// TIA Portal project "S7_1516_LECTOR620_DI" (V15)

(* hardware
DEVICE "S71500/ET200MP station_1"  S7-1500 station
   slot 0: "Rail_0"  Rack  6ES7 590-1***0-0AA0
   slot 0: "PM 190W 120/230VAC"  PM 190W 120/230VAC  6EP1333-4BA00
   slot 1: "PLC_1"  CPU 1516-3 PN/DP  6ES7 516-3AN00-0AB0  V1.8
      slot 3: "CPU display_1"  6ES7591-1BA00-0AA0
   slot 2: "DI 32x24VDC HF_1"  DI 32x24VDC HF  6ES7 521-1BL00-0AB0  V2.1
   slot 3: "DQ 32x24VDC/0.5A ST_1"  DQ 32x24VDC/0.5A ST  6ES7 522-1BL00-0AB0  V2.0
   slot 4: "AI 8xU/I/RTD/TC ST_1"  AI 8xU/I/RTD/TC ST  6ES7 531-7KF00-0AB0  V2.0
   slot 5: "AQ 4xU/I ST_1"  AQ 4xU/I ST  6ES7 532-5HD00-0AB0  V2.0
DEVICE "HMI_1"  TP700 Comfort
   slot 0: "HMI_1"  TP700 Comfort  6AV2 124-0GC01-0AX0  15.0.0.0
   slot 1: "HMI_RT_1"  TP700 Comfort  6AV2 124-0GC01-0AX0  15.0.0.0
   slot 5: "HMI_1.IE_CP_1"  PROFINET Interface  15.0.0.0
      slot 1: "PROFINET Interface_1"  PROFINET Interface
         slot 1: "Port_1"  Port
         slot 2: "Port_2"  Port
   slot 7: "HMI_1.MPI/DP_CP_1"  MPI/DP Interface  15.0.0.0
DEVICE "GSD device_2"  GSD.Device.PN
   slot 0: "Rack"  Rack  V1.0
   slot 0: "LECTOR62x"  LECTOR62x  HandShake (HS)  V1.1.0
      slot 0: "LECTOR62x  HandShake (HS)"  LECTOR62x  HandShake (HS)
      slot 1: "Interface"  Interface
         slot 1: "Port 1"  Port 1
   slot 1: "Ctrl Bits in_1"  Ctrl Bits in
      slot 0: "Ctrl Bits in"  Ctrl Bits in
   slot 2: "Ctrl Bits out_1"  Ctrl Bits out
      slot 0: "Ctrl Bits out"  Ctrl Bits out
   slot 3: " 32 Byte Input (HS)_1"   32 Byte Input (HS)
      slot 0: " 32 Byte Input (HS)"   32 Byte Input (HS)
   slot 4: " 32 Byte Output (HS)_1"   32 Byte Output (HS)
      slot 0: " 32 Byte Output (HS)"   32 Byte Output (HS)
DEVICE "PC-System_1"  SIMATIC PC station
   slot 0: "SIMATIC PC station"  Rail  SIMATIC PC-Station  V1.0
      slot 125: "Stationmanager"  Station_Manager  V6.0.4
   slot 1: "IE general_1"  IE General  IE_CP  V8.2.0
   slot 3: "HMI_RT_2"  WinCC RT Advanced  6AV2 104-0xxxx-xxxx  15.0.0.0
      slot 33792: "Host interface"  Host interface
*)

// ===== PLC "PLC_1"  CPU 1516-3 PN/DP =====

VAR_GLOBAL   // PLC tag table "Default tag table"
   "AD_CH0" AT %IW4 : Int;
   "Sensor1" AT %I0.0 : Bool;
   "Tag_5" AT %IW58 : Int;
   "Tag_6" AT %IW12 : Int;
   "DA_CH0" AT %QW4 : Int;
   "SICK_IN_1" AT %Q0.0 : Bool;
   "Tag_3" AT %Q0.1 : Bool;
   "Tag_4" AT %QW1 : Int;
   "Tag_7" AT %Q0.2 : Bool;
   "Tag_8" AT %Q1.1 : Bool;
   "Tag_9" AT %Q1.2 : Bool;
   "Clock_Byte" AT %MB0 : Byte;
   "Clock_10Hz" AT %M0.0 : Bool;
   "Clock_5Hz" AT %M0.1 : Bool;
   "Clock_2.5Hz" AT %M0.2 : Bool;
   "Clock_2Hz" AT %M0.3 : Bool;
   "Clock_1.25Hz" AT %M0.4 : Bool;
   "Clock_1Hz" AT %M0.5 : Bool;
   "Clock_0.625Hz" AT %M0.6 : Bool;
   "Clock_0.5Hz" AT %M0.7 : Bool;
   "SignalUlaz" AT %M1.0 : Bool;
   "SICK_OUT_1" AT %I0.1 : Bool;
   "SICK_OUT_1_MEM" AT %M10.0 : Bool;
   "Tag_1" AT %M100.0 : Bool;
   "Tag_2" AT %M100.1 : Bool;
   "Tag_10" AT %M100.2 : Bool;
   "Tag_11" AT %M100.3 : Bool;
   "Tag_12" AT %MW101 : Word;
   "Request" AT %M100.4 : Bool;
   "No_of_counts_in" AT %IB57 : Byte;
   "No_of_counts_out" AT %QB49 : Byte;
   "SICK_OUT_1_old" AT %M2.0 : Bool;
   "Code_byte_1" AT %IB62 : Byte;
   "Tag_13" AT %MW3 : Int;
   "MOVE_ERROR" AT %MW4 : Int;
   "Tag_14" AT %IB56 : Byte;
   "Code_byte_2" AT %IB63 : Char;
   "Code_byte_3" AT %IB64 : Char;
   "Code_byte_4" AT %IB65 : Char;
   "Code_byte_5" AT %IB66 : Char;
   "Code_byte_6" AT %IB67 : Char;
   "Code_byte_7" AT %IB68 : Char;
   "Code_byte_8" AT %IB69 : Char;
   "Code_byte_9" AT %IB70 : Char;
   "Code_byte_10" AT %IB71 : Char;
   "Code_byte_11" AT %IB72 : Char;
   "Code_byte_12" AT %IB73 : Char;
   "Code_byte_13" AT %IB74 : Char;
   "ADDA_ENABLE" AT %I0.2 : Bool;
   "DA_CH2" AT %QW8 : Int;
   "AD_CH2" AT %IW8 : Int;
   "AD_CH1" AT %IW6 : Int;
   "AD_CH3" AT %IW10 : Int;
   "DA_CH1" AT %QW6 : Int;
   "DA_CH3" AT %QW10 : Int;
   "iCounter_Tag_kopija" AT %QW12 : Int;
   "PrebranaKoda" AT %QW14 : WChar;
   "Tag_15" AT %I0.3 : Bool;
   "Tag_16" AT %Q0.3 : Bool;
   "Tag_17" AT %Q2.0 : Bool;
   "Tag_18" AT %Q2.1 : Bool;
   "Tag_19" AT %Q2.2 : Bool;
END_VAR

// folder: SICK AG

TYPE "ST_SICK_Lector_CLV6xx"
TITLE = SICK Lector/CLV6xx data type
VERSION : 0.1
// This data type includes arguments and results using by the SICK_Lector_CLV6xx_PNDP function block.
   STRUCT
      Matchcode : Struct   // ==Matchcode==
         sName : String[10];   // Matchcode number (Match[1..9]) (Input)
         nCodeType : Char;   // Code type see device documentation. (Example: 'd'= EAN-Code; 's'=QR-Code; '*'= Don't care) (Input)
         iMinMaxLength : USInt;   // Sets the min and may length. 0= Don't care (Input)
         sContent : String[75];   // Matchcode content
      END_STRUCT;
      FreeCommand : Struct   // ==Free Command==
         sCommand : String[100];   // Command (SICK CoLa-A protocol without [STX]/[ETX] framing) (In)
         sResult : String[100];   // Result (SICK CoLa-A protocol) (Out)
      END_STRUCT;
      ReadingResult : Struct   // ==Reading Result==
         iCounter : USInt;   // This counter is incremented if a new reading result has arrived (In)
         iLength : Int;   // Byte length of the reading result (Out)
         arrResult : Array[1..200] of Byte;   // Reading result data defined in the SOPAS output format (Out)
      END_STRUCT;
   END_STRUCT;
END_TYPE

// folder: (top level)

DATA_BLOCK "Data_block_1"   // DB1
{ S7_Optimized_Access := 'FALSE' }
VERSION : 0.1
   VAR
      Error_Detektovan : Bool;   // 1 ce je prislo do napake
      Error_Koda : DWord;   // ID koda napake
      startFound : Bool;   // za Move_Code funkcijo
      endFound : Bool;   // za Move_Code funkcijo
      Sensor_ok_blink : Byte;
      No_of_counts : LInt;
      DA0 : Real;
      AD0 : Real;
      DA2 : Real;
      AD2 : Real;
      Static_1 : Array[0..5] of Int;
      TestBitStefanRequest : Bool;
      ShranjenaPrebranaKoda_Cas : Date_And_Time := DT#2021-05-14-08:00:42.263;
      ShranjenaPrebranaKoda : String;
      Operand1 : Bool;
      DatumInCas : Struct
         Datum : Bool;
         Ura : Bool;
      END_STRUCT;
      AD3 : Real;
      Prebrana_Koda_FLAG : Bool;
      Counter_1_Reset : Bool;
      Operand2 : Bool;
   END_VAR
BEGIN
END_DATA_BLOCK

DATA_BLOCK "IDB_Lector6xx"   // DB2
{ S7_Optimized_Access := 'TRUE' }
AUTHOR : SICKAG
FAMILY : Ident
VERSION : 1.2
// stored: InstanceOfName SICK_Lector_CLV6xx_PNDP
"SICK_Lector_CLV6xx_PNDP"
BEGIN
END_DATA_BLOCK

DATA_BLOCK "DB_Example"   // DB3
{ S7_Optimized_Access := 'TRUE' }
VERSION : 0.1
   VAR
      stEdge : Struct   // Edge detection flags
         xEdgeTrigger : Bool;
         xEdgeMatchcode : Bool;
         xEdgeDone : Bool;
         xEdgeError : Bool;
         xEdgeTriggerMem : Bool;
         xEdgeDoneMem : Bool;
         xEdgeErrorMem : Bool;
         xEdgeMatchcodeMem : Bool;
      END_STRUCT;
      xTrigger : Bool;   // Start read tag command
      xMatchcode : Bool;
      xTriggerDone : Bool;   // Read tag done
      xMatchcodeDone : Bool;
      sReadingResult : String[200];   // Read content
      stLector : "ST_SICK_Lector_CLV6xx";   // RFU data
      arrReadingResult : Array[0..199] of Byte;   // Read content backup
   END_VAR
BEGIN
END_DATA_BLOCK

DATA_BLOCK "SICK_Lector_CLV6xx_PNDP_DB"   // DB4
{ S7_Optimized_Access := 'TRUE' }
AUTHOR : SICKAG
FAMILY : Ident
VERSION : 1.2
// stored: InstanceOfName SICK_Lector_CLV6xx_PNDP
"SICK_Lector_CLV6xx_PNDP"
BEGIN
END_DATA_BLOCK

DATA_BLOCK "Block_1_DB"   // DB5
{ S7_Optimized_Access := 'TRUE' }
AUTHOR : Stefan_Milivojcev
VERSION : 0.1
// stored: InstanceOfName Block_1
"Block_1"
BEGIN
END_DATA_BLOCK

// folder: System blocks/Program resources

DATA_BLOCK "IEC_Counter_0_DB"   // DB6
{ S7_Optimized_Access := 'TRUE' }
AUTHOR : SIMATIC
FAMILY : IEC
NAME : LCNTR
VERSION : 1.2
// stored: InstanceOfName IEC_LCOUNTER
"IEC_LCOUNTER"
BEGIN
END_DATA_BLOCK

// folder: (top level)

FUNCTION_BLOCK "Block_1"   // FB1, SCL
TITLE = Shranjevanje_Branja
{ S7_Optimized_Access := 'TRUE' }
AUTHOR : Stefan_Milivojcev
VERSION : 0.1
   VAR_INPUT
      RESULT_ARRAY_SIZE : Int;   // Velikost najvecjega moznega rezultata branja
      Date_Time_Temp : Date_And_Time;
   END_VAR
   VAR_OUTPUT
      startFound : Bool;
      endFound : Bool;
      PrebranaKoda_Cas : Date_And_Time;
      PrebranaKoda : String;
   END_VAR
   VAR_TEMP
      i : Int;
   END_VAR
BEGIN
   //Stefan Milivojčev
   //stefan.milivojcev@gmail.com
   //
   //Prepoznava START in STOP bita


   #startFound := FALSE;
   #endFound := FALSE;
   #i := 0;
   #PrebranaKoda := '';



   IF ("DB_Example".stLector.ReadingResult.arrResult[1] = 16#02) THEN
       // Statement section IF
       #startFound := 1;
   END_IF;

   IF (#startFound = 1) THEN //ce smo najdli zacetek kode iscemo konec

       FOR #i := 1 TO #RESULT_ARRAY_SIZE DO
           // Statement section FOR

           IF ("DB_Example".stLector.ReadingResult.arrResult[#i] = 16#03) THEN
               // Statement section IF
               #endFound := TRUE;

           ELSE

               #PrebranaKoda[#i - 1] := "DB_Example".stLector.ReadingResult.arrResult[#i];

           END_IF;



       END_FOR;

       #PrebranaKoda_Cas := #Date_Time_Temp;


   END_IF;




   "Data_block_1".No_of_counts := "DB_Example".stLector.ReadingResult.iCounter;
END_FUNCTION_BLOCK

ORGANIZATION_BLOCK "Main"   // OB1, LAD, ProgramCycle
TITLE = "Main Program Sweep (Cycle)"
{ S7_Optimized_Access := 'TRUE' }
VERSION : 0.1
   VAR_INPUT
      Initial_Call : Bool;   // Initial call of this OB
      Remanence : Bool;   // =True, if remanent data are available
   END_VAR
   VAR_TEMP
      Temp_3 : Real;
      Temp_2 : LInt;
      Temp_Cas_Branja : Date_And_Time;
      Temp3 : Date;
      Temp4 : DInt;
      temp6 : Bool;
      Temp5 : UInt;
   END_VAR
   VAR_TEMP   // added for the SCL form of the ladder/FBD networks
      _w1 : Bool;
      _w2 : Bool;
   END_VAR
BEGIN

REGION Network 1: Request za branje
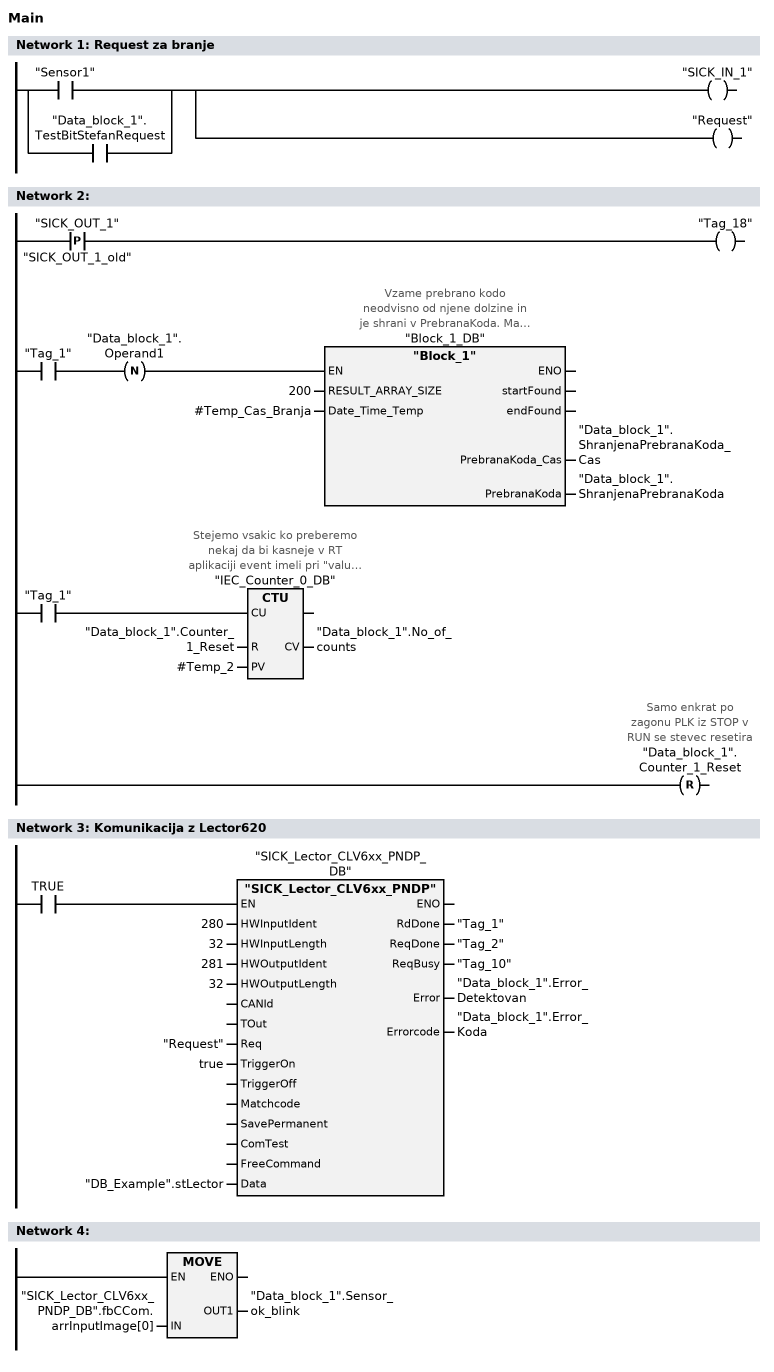
   RUNG wire#powerrail
      Contact( "Sensor1" )
      wire#w1
      Coil( "SICK_IN_1" )
   END_RUNG
   RUNG wire#powerrail
      Contact( "Data_block_1".TestBitStefanRequest )
   END_RUNG wire#w1
   RUNG wire#w1
      Coil( "Request" )
   END_RUNG
   // the same network as SCL:
   "SICK_IN_1" := "Sensor1" OR "Data_block_1".TestBitStefanRequest;
   "Request" := "SICK_IN_1";
END_REGION

REGION Network 2
   #_w1 := "SICK_OUT_1" AND NOT "SICK_OUT_1_old";   // rising edge of "SICK_OUT_1"
   "SICK_OUT_1_old" := "SICK_OUT_1";
   "Tag_18" := #_w1;
   #_w2 := NOT "Tag_1" AND "Data_block_1".Operand1;   // falling edge
   "Data_block_1".Operand1 := "Tag_1";
   IF #_w2 THEN
       "Block_1_DB"(RESULT_ARRAY_SIZE := 200,   // "Block_1": Vzame prebrano kodo neodvisno od njene dolzine in je shrani v PrebranaKoda. Max dolzina je trenutno 200
                    Date_Time_Temp := #Temp_Cas_Branja,
                    PrebranaKoda_Cas => "Data_block_1".ShranjenaPrebranaKoda_Cas,
                    PrebranaKoda => "Data_block_1".ShranjenaPrebranaKoda);
   END_IF;
   "IEC_Counter_0_DB".CTU(CU := "Tag_1",   // Stejemo vsakic ko preberemo nekaj da bi kasneje v RT aplikaciji event imeli pri "value change"
                          R := "Data_block_1".Counter_1_Reset,
                          PV := #Temp_2,
                          CV => "Data_block_1".No_of_counts);
   "Data_block_1".Counter_1_Reset := FALSE;   // Samo enkrat po zagonu PLK iz STOP v RUN se stevec resetira
END_REGION

REGION Network 3: Komunikacija z Lector620
   RUNG wire#powerrail
      Contact( TRUE )
      "SICK_Lector_CLV6xx_PNDP_DB"(HWInputIdent := 280, HWInputLength := 32, HWOutputIdent := 281, HWOutputLength := 32, CANId :=, TOut :=, Req := "Request", TriggerOn := true, TriggerOff :=, Matchcode :=, SavePermanent :=, ComTest :=, FreeCommand :=, Data := "DB_Example".stLector, RdDone => "Tag_1", ReqDone => "Tag_2", ReqBusy => "Tag_10", Error => "Data_block_1".Error_Detektovan, Errorcode => "Data_block_1".Error_Koda)
   END_RUNG
   // the same network as SCL:
   IF TRUE THEN
       "SICK_Lector_CLV6xx_PNDP_DB"(HWInputIdent := 280,   // "SICK_Lector_CLV6xx_PNDP"
                               HWInputLength := 32,
                               HWOutputIdent := 281,
                               HWOutputLength := 32,
                               Req := "Request",
                               TriggerOn := true,
                               Data := "DB_Example".stLector,
                               RdDone => "Tag_1",
                               ReqDone => "Tag_2",
                               ReqBusy => "Tag_10",
                               Error => "Data_block_1".Error_Detektovan,
                               Errorcode => "Data_block_1".Error_Koda);
   END_IF;
END_REGION

REGION Network 4
   RUNG wire#powerrail
      Move(in := "SICK_Lector_CLV6xx_PNDP_DB".fbCCom.arrInputImage[0], out1 => "Data_block_1".Sensor_ok_blink)
   END_RUNG
   // the same network as SCL:
   "Data_block_1".Sensor_ok_blink := "SICK_Lector_CLV6xx_PNDP_DB".fbCCom.arrInputImage[0];
END_REGION
END_ORGANIZATION_BLOCK

ORGANIZATION_BLOCK "Cyclic interrupt"   // OB30, LAD, CyclicInterrupt
{ S7_Optimized_Access := 'TRUE' }
VERSION : 0.1
   VAR_INPUT
      Initial_Call : Bool;   // Initial call of this OB
      Event_Count : Int;   // Events discarded
   END_VAR
BEGIN

REGION Network 1
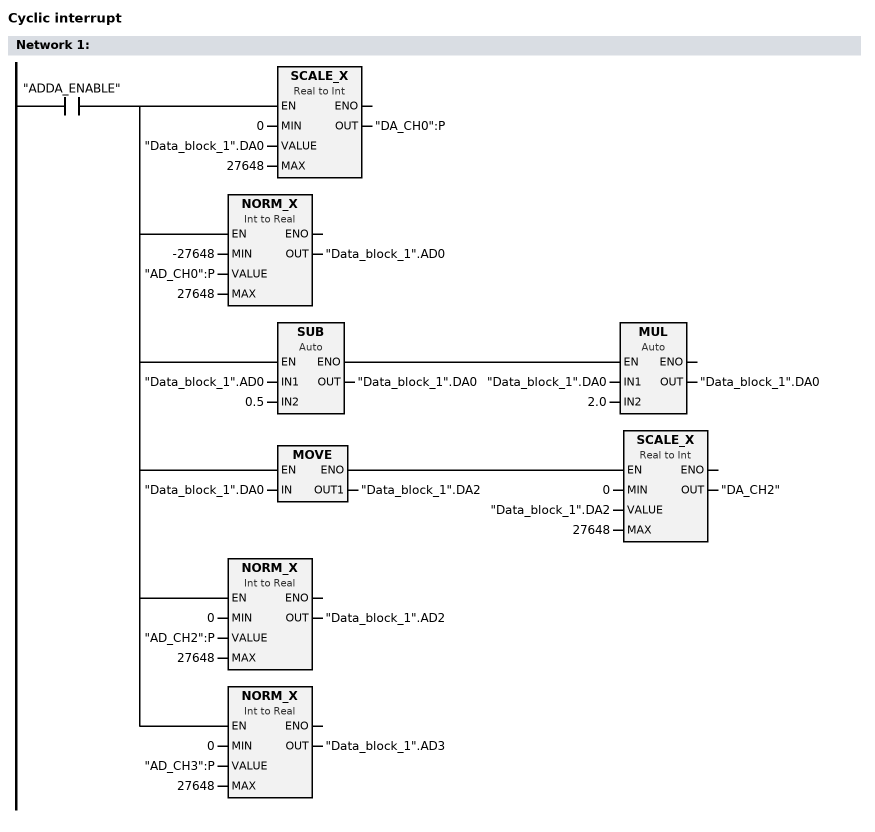
   RUNG wire#powerrail
      Contact( "ADDA_ENABLE" )
      wire#w1
      { S7_Templates := "[SrcType := Real, DestType := Int]" } Scale(min := 0, value := "Data_block_1".DA0, max := 27648, out => "DA_CH0":P)
   END_RUNG
   RUNG wire#w1
      { S7_Templates := "[SrcType := Int, DestType := Real]" } Normalize(min := -27648, value := "AD_CH0":P, max := 27648, out => "Data_block_1".AD0)
   END_RUNG
   RUNG wire#w1
      Sub(in1 := "Data_block_1".AD0, in2 := 0.5, out => "Data_block_1".DA0)
      Mul(in1 := "Data_block_1".DA0, in2 := 2.0, out => "Data_block_1".DA0)
   END_RUNG
   RUNG wire#w1
      Move(in := "Data_block_1".DA0, out1 => "Data_block_1".DA2)
      { S7_Templates := "[SrcType := Real, DestType := Int]" } Scale(min := 0, value := "Data_block_1".DA2, max := 27648, out => "DA_CH2")
   END_RUNG
   RUNG wire#w1
      { S7_Templates := "[SrcType := Int, DestType := Real]" } Normalize(min := 0, value := "AD_CH2":P, max := 27648, out => "Data_block_1".AD2)
   END_RUNG
   RUNG wire#w1
      { S7_Templates := "[SrcType := Int, DestType := Real]" } Normalize(min := 0, value := "AD_CH3":P, max := 27648, out => "Data_block_1".AD3)
   END_RUNG
   // the same network as SCL:
   IF "ADDA_ENABLE" THEN
       "DA_CH0":P := SCALE_X(MIN := 0, VALUE := "Data_block_1".DA0, MAX := 27648);
       "Data_block_1".AD0 := NORM_X(MIN := -27648, VALUE := "AD_CH0":P, MAX := 27648);
       "Data_block_1".DA0 := "Data_block_1".AD0 - 0.5;
       "Data_block_1".DA0 := "Data_block_1".DA0 * 2.0;
       "Data_block_1".DA2 := "Data_block_1".DA0;
       "DA_CH2" := SCALE_X(MIN := 0, VALUE := "Data_block_1".DA2, MAX := 27648);
       "Data_block_1".AD2 := NORM_X(MIN := 0, VALUE := "AD_CH2":P, MAX := 27648);
       "Data_block_1".AD3 := NORM_X(MIN := 0, VALUE := "AD_CH3":P, MAX := 27648);
   END_IF;
END_REGION
END_ORGANIZATION_BLOCK

ORGANIZATION_BLOCK "Startup"   // OB100, LAD, Startup
TITLE = "Complete Restart"
{ S7_Optimized_Access := 'TRUE' }
VERSION : 0.1
   VAR_INPUT
      LostRetentive : Bool;   // True if retentive data are lost
      LostRTC : Bool;   // True if date and time are lost
   END_VAR
   VAR_TEMP
      operand1 : Bool;
   END_VAR
BEGIN

REGION Network 1
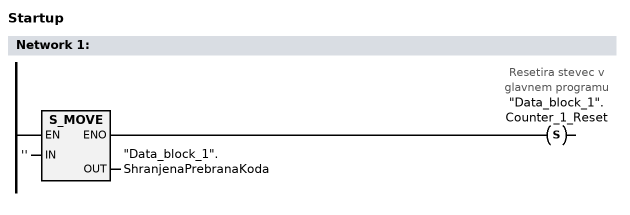
   RUNG wire#powerrail
      S_Move(in := '', out => "Data_block_1".ShranjenaPrebranaKoda)
      S_Coil( "Data_block_1".Counter_1_Reset )   // Resetira stevec v glavnem programu
   END_RUNG
   // the same network as SCL:
   "Data_block_1".ShranjenaPrebranaKoda := '';
   "Data_block_1".Counter_1_Reset := TRUE;   // Resetira stevec v glavnem programu
END_REGION
END_ORGANIZATION_BLOCK

// folder: SICK AG

FUNCTION_BLOCK "SICK_Lector_CLV6xx_PNDP"   // FB72, SCL
TITLE = SICK Lector6xx / CLV6xx function block
{ S7_Optimized_Access := 'TRUE' }
AUTHOR : SICKAG
FAMILY : Ident
VERSION : 1.2
// This function block is used for a communication between a SICK Lector6xx / SICK CLV6xx code reader and a Siemens S7-1200/S7-1500 PLC via  PROFINET/PROFIBUS
   VAR_INPUT
      HWInputIdent : Hw_Io;   // Hardware identification number of the input module
      HWInputLength : USInt;   // Size of the input module
      HWOutputIdent : Hw_Io;   // Hardware identification number of the output module
      HWOutputLength : USInt;   // Size of the output module
      CANId : USInt;   // CAN ID (0= Master / No CAN network)
      TOut : Time := T#10s;   // Time out
      Req : Bool;   // A positive edge starts the request
      TriggerOn : Bool;   // Select: Trigger On to open the reading gate via a SW-Trigger command
      TriggerOff : Bool;   // Select: Trigger Off to close the reading gate via a SW-Trigger command
      Matchcode : Bool;   // Select: Matchcode (details at #Data)
      SavePermanent : Bool;   // Select: Save permanent
      ComTest : Bool;   // Select: Communication test
      FreeCommand : Bool;   // Select: Free command (details at #Data)
   END_VAR
   VAR_OUTPUT
      RdDone : Bool;   // Positive edge: A reading result sent by the device was received
      ReqDone : Bool;   // Request done / Indicates whether a CoLa command was sent and an answer was received
      ReqBusy : Bool;   // Request in process / Request processing
      Error : Bool;   // Error detected
      Errorcode : DWord;   // Error code (see documentation)
   END_VAR
   VAR_IN_OUT
      Data : "ST_SICK_Lector_CLV6xx";   // Command arguments and result outputs of the FB actions
   END_VAR
   VAR
      bTriggerReq : Bool;   // Rising edge detection
      bTriggerReqMem : Bool;   // Rising edge detection
      bTriggerDone : Bool;   // Rising edge detection
      bTriggerDoneMem : Bool;   // Rising edge detection
      bTriggerError : Bool;   // Rising edge detection
      bTriggerErrorMem : Bool;   // Rising edge detection
      bCanActive : Bool;   // CAN-Bus active flag
      bDeviceState : Bool;   // Current device state (True= Edit-Mode | False= Run-Mode)
      bEnforceLogout : Bool;   // Logout enforced
      bReqBusyMem : Bool;   // Backup variable
      iStep : USInt;   // Currrent FB step
      iCommandIndex : Int;   // Command index
      iCommandLength : UInt;   // Length of the command that should be send
      iRecordSize : UInt;   // Length of the record array
      iCommandSize : UInt;   // Length of the command array
      iReadingResultSize : UInt;   // Length of the reading result array
      iIndex : UInt;   // Index variable
      nTempErrorCode : DWord;   // Temporarily error code
      nLogoutErrorCode : DWord;   // Temporarily error code
      arrSelection : Array[0..5] of Bool;   // input bit selection
      arrCommand : Array[0..499] of Byte;   // Contains the transmitted CoLa command
      arrRecord : Array[0..499] of Byte;   // Contains the received telegram
      fbTimeout : TON_TIME;   // Instance: Timer on delay (Time out)
      fbCCom : "SICK_CCOMM_PNDP";   // Instance: CoLa communication block
   END_VAR
   VAR_TEMP
      iTemp1 : Int;   // Temporarily variable
      iTemp2 : UDInt;   // Temporarily variable
      iTemp3 : UDInt;   // Temporarily variable
      nFncValue : DWord;   // Get/Set function value
      nFncErrorCode : Word;   // Get/Set function error code
   END_VAR
BEGIN
   (*===========================================================================================
   Name:   SICK_Lector_CLV6xx_PNDP 
   Author: SICK AG
   =============================================================================================
   Description: 
   This function block is used for a communication between a SICK Lector6xx / SICK CLV6xx
   code reader and a Siemens S7-1200/S7-1500 PLC via PROFINET/PROFIBUS.                         

   =============================================================================================
   Features:        
   - Receive reading results of the device, triggered by a command, fieldbus or by a hardware 
     switch. The content of the result can be modified in the "Output Format" option in the
     SOPAS engineeringtool.                                           
   - Open and close a reading gate (software trigger via command)
   - Set a new Matchcode evaluation condition 
   - Save all device parameters permanent                                                  
   - Communication test
   - Send a free defined CoLa-A telegram and receive the result
   - All commands can also be used in a SICK CAN-Bus network

   =============================================================================================
   Version history:
   Date       | Version | Author  | Remark
   ---------------------------------------------------------------------------------------------
   21/02/2014 | V1.0    | SICK AG | Initial version
   07/08/2014 | V1.1    | SICK AG | Replace R_TRIG function 
   24/10/2017 | V1.2    | SICK AG | Avoid initialization warnings which occurs using TIA V13 or higher
   ============================================================================================*)

   (*===================================== INITIALISATION =====================================*)
   #iRecordSize:= 500;         (*Length of the arrRecord array*)
   #iCommandSize:= 500;        (*Length of the arrCommand array*)
   #iReadingResultSize:= 200;  (*Length of the reading result array*)

   (*Rising edge detection*)
   #bTriggerReq:= #Req AND NOT #bTriggerReqMem;
   #bTriggerReqMem:= #Req;
   #bTriggerDone:= #fbCCom.ReqDone AND NOT #bTriggerDoneMem;
   #bTriggerDoneMem:= #fbCCom.ReqDone;
   #bTriggerError:= #fbCCom.Error AND NOT #bTriggerErrorMem;
   #bTriggerErrorMem:= #fbCCom.Error;

   (*Reset the read done flag every cycle*)
   #RdDone:= false;


   (*===================================== ERROR HANDLING =====================================*)
   (* bDeviceState  |  bEnforceLogout  |  Action
          FALSE     |      FALSE       |  Errorcode = Errorcode from last plc cycle
          FALSE     |      TRUE        |  Errorcode = Logout error
          TRUE      |      FALSE       |  Enforce "Logout" command
          TRUE      |      TRUE        |  Errorcode = Logout not possible + Reason*)
   IF #nTempErrorCode <>16#0000_0000 THEN

     (*Enfore "Logout" command*)
     IF #bDeviceState AND NOT #bEnforceLogout THEN
       #bEnforceLogout:= true;
       #iCommandIndex:= 11;                  (*Logout*)
       #nLogoutErrorCode:= #nTempErrorCode;  (*Save current error code*)
       #nTempErrorCode:= 16#0000_0000;       (*Clear currenr error variable*)
       #iStep:= 4;                           (*Create command*)

     (*Logout can not be ensured*)
     ELSIF #bDeviceState AND #bEnforceLogout THEN
       #Errorcode.%W1:= #nTempErrorCode.%W0;  
       #Errorcode.%W0:= 16#0017;  (*Error: Logout can not be ensured (please check the device state)*)

     (*Errorcode = Errorcode from the last plc cycle or logout error*)
     ELSE
       #Errorcode:= #nTempErrorCode;
     END_IF;

     (*Update FB status*)
     IF #nTempErrorCode <> 16#0000_0000 THEN
       #ReqDone:= false;
       #ReqBusy:= false;
       #bReqBusyMem:= false;
       #Error:= true;
       #nTempErrorCode:= 16#0000_0000;
       #nLogoutErrorCode:= 16#0000_0000;
       #iStep:= 0;
       RETURN;
     END_IF;
   END_IF;

   (*Time out detection*)
   #fbTimeout(IN:= #bReqBusyMem, PT:= #TOut);
   IF #fbTimeout.Q THEN
     #nTempErrorCode:= 16#0000_0010; (*Error: Time out*)
   END_IF;

   (*Check if a device error is detected: 'sFA XX'*)
   IF #bTriggerDone AND ((NOT #bCanActive AND
     #arrRecord[0] = 's' AND
     #arrRecord[1] = 'F' AND
     #arrRecord[2] = 'A') OR (#bCanActive AND
     #arrRecord[0] = 's' AND
     #arrRecord[12] = 'F' AND
     #arrRecord[13] = 'A')) THEN

     (*Get the position of the error code*)
     IF #bCanActive THEN
       #iIndex:= 15;
     ELSE
       #iIndex:= 4;
     END_IF;

     "SICK_GetValue"(iTelegramLength:= INT_TO_UINT(#fbCCom.ReqLength),
                     iValueLength:= 0,
                     nValue=> #nFncValue,
                     nErrorCode=> #nFncErrorCode,
                     iPosition:= #iIndex,
                     arrData:= #arrRecord);

     IF #nFncErrorCode = 16#0000 THEN
       #nTempErrorCode.%W1:= DWORD_TO_WORD(#nFncValue);
       #nTempErrorCode.%W0:= 16#0011; (*Error: Device error*)
     ELSE
       #nTempErrorCode.%W1:= #nFncErrorCode;
       #nTempErrorCode.%W0:= 16#0012; (*Error: SICK_GetValue error*)      
     END_IF;
   END_IF;

   (*Error detected*)
   IF #nTempErrorCode <>16#0000_0000 THEN
     RETURN;
   END_IF;


   (*================================= START REQUEST (STEP 1) =================================*)
   IF NOT #bReqBusyMem AND #bTriggerReq THEN
     #ReqDone:= false;
     #ReqBusy:= true;
     #bReqBusyMem:= true;
     #Error:= false;
     #Errorcode:= 16#0000_0000;
     #bDeviceState:= false;
     #bEnforceLogout:= false;

     (*Save the current bit selection for the job*)
     #arrSelection[0]:= #TriggerOn;
     #arrSelection[1]:= #TriggerOff;
     #arrSelection[2]:= #Matchcode;
     #arrSelection[3]:= #SavePermanent;
     #arrSelection[4]:= #ComTest;
     #arrSelection[5]:= #FreeCommand;


     (*Check CAN-ID*)
     IF #CANId > 63 THEN
       #nTempErrorCode:= 16#0000_0014; (*Error invalid CAN Id*)  
     ELSIF #CANId = 0 THEN
       #bCanActive:= false;
       #iStep:= 3; (*Check parameter input*)
     ELSE
       #bCanActive:= true;
       #iStep:= 2; (*Add CAN identifier*)
     END_IF;
   END_IF;


   (*=============================== ADD CAN IDENTIFIER (STEP 2) ==============================*)
   IF #iStep =2 THEN
     Strg_TO_Chars(Strg:= 's{ 00 01 ', pChars:= 0, Cnt=> #iIndex, Chars:=#arrCommand);

     "SICK_SetValue"(bAddBlank:= false,
                     nValue:= #CANId,
                     arrData=> #arrCommand,
                     nErrorCode=> #nFncErrorCode,
                     iPosition:= #iIndex);
     IF #nFncErrorCode <> 16#0000 THEN
       #nTempErrorCode.%W1:= #nFncErrorCode;
       #nTempErrorCode.%W0:= 16#0013; (*Error: SICK_SetValue error*)
     ELSE
       #arrCommand[#iIndex]:= '}';
       #iStep:= 3; (*Check parameter input*)
     END_IF;
   END_IF;


   (*============================= CHECK PARAMETER INPUT (STEP 3) =============================*)
   IF #iStep =3 THEN
     #iTemp1:= 0; (*Counts up the active bit selection*)

     (*Command: Trigger On*)
     IF #arrSelection[0] THEN
       #iTemp1:= #iTemp1+1;
       #iCommandIndex:= 0; (*Send a "Trigger On" command*)
     END_IF;

     (*Command: Trigger Off*)
     IF #arrSelection[1] THEN
       #iTemp1:= #iTemp1+1;
       #iCommandIndex:= 1; (*Send a "Trigger Off" command*)
     END_IF;

     (*Command: Matchcode*)
     IF #arrSelection[2] THEN
       #iTemp1:= #iTemp1+1;

       IF #Data.Matchcode.sName = '' THEN
         #nTempErrorCode:= 16#0000_0022; (*Error: Matchcode name is empty*)
       ELSIF #Data.Matchcode.nCodeType <='$20' OR #Data.Matchcode.nCodeType > '$7E' THEN
         #nTempErrorCode:= 16#0000_0023; (*Error: Invalid code type*)
       END_IF;

       #iCommandIndex:= 10; (*Send a "Login" command*)
     END_IF;

     (*Command: Save permanent*)
     IF #arrSelection[3] THEN 
       #iTemp1:= #iTemp1+1;
       #iCommandIndex:= 10; (*Send a "Login" command*)  
     END_IF;

     (*Command: Communication test*)
     IF #arrSelection[4] THEN
       #iTemp1:= #iTemp1+1;
       #iCommandIndex:= 4; (*Send a "Comm Test" command*)
     END_IF;

     (*Command: Free command*)
     IF #arrSelection[5] THEN
       #iTemp1:= #iTemp1+1;

       (*Check length*)
       IF #bCanActive THEN
         #iTemp2:= INT_TO_UDINT(LEN(#Data.FreeCommand.sCommand))+11;
       ELSE
         #iTemp2:= INT_TO_UDINT(LEN(#Data.FreeCommand.sCommand));
       END_IF;

       IF (LEN(#Data.FreeCommand.sCommand) <=0) OR (#iTemp2 > #iCommandSize) THEN
         #nTempErrorCode:= 16#0000_0020; (*Error: Invalid free command length*)
       END_IF;

       #iCommandIndex:= 5; (*Send a "Free Command" command*)
     END_IF;

     (*Check bit sum of the command selection*)
     IF #iTemp1 <>1 THEN
       #nTempErrorCode:= 16#0000_0015; (*Error: More than one or no parameter selected*)   
     END_IF;

     (*Check if a error was detected*)
     IF #nTempErrorCode = 16#0000_0000 THEN
       #iStep:= 4; (*Create CoLa command*)
     END_IF;
   END_IF;


   (*============================== CREATE COLA COMMAND (STEP 4) ==============================*)
   IF #iStep =4 THEN
     CASE #iCommandIndex OF

     (*Create "Trigger On" command*)
     0:  IF #bCanActive THEN
           Strg_TO_Chars(Strg:= 'MN mTCgateon', pChars:= 12, Cnt=> #iTemp3, Chars:=#arrCommand);
           #iCommandLength:= UDINT_TO_UINT(#iTemp3)+12;
         ELSE
           Strg_TO_Chars(Strg:= 'sMN mTCgateon', pChars:= 0, Cnt=> #iTemp3, Chars:=#arrCommand);
           #iCommandLength:= UDINT_TO_UINT(#iTemp3);
         END_IF;
         #iStep:= 5; (*Send command*)

     (*Create "Trigger Off" command*)
     1:  IF #bCanActive THEN
           Strg_TO_Chars(Strg:= 'MN mTCgateoff', pChars:= 12, Cnt=> #iTemp3, Chars:=#arrCommand);
           #iCommandLength:= UDINT_TO_UINT(#iTemp3)+12;
         ELSE
           Strg_TO_Chars(Strg:= 'sMN mTCgateoff', pChars:= 0, Cnt=> #iTemp3, Chars:=#arrCommand);
           #iCommandLength:= UDINT_TO_UINT(#iTemp3);
         END_IF;
         #iStep:= 5; (*Send command*)

     (*Create "Matchcode" command*)
     2:  IF #bCanActive THEN
           Strg_TO_Chars(Strg:= 'MN mEVSetMatchCode 00 ', pChars:= 12, Cnt=> #iTemp3, Chars:=#arrCommand);
           #iIndex:= UDINT_TO_UINT(#iTemp3+12);
         ELSE
           Strg_TO_Chars(Strg:= 'sMN mEVSetMatchCode 00 ', pChars:= 0, Cnt=> #iTemp3, Chars:=#arrCommand);
           #iIndex:= UDINT_TO_UINT(#iTemp3);
         END_IF;

         (*Add matchcode name*)
         Strg_TO_Chars(Strg:= CONCAT(IN1:= 'name="', IN2:= #Data.Matchcode.sName), pChars:= #iIndex, Cnt=> #iTemp3, Chars:=#arrCommand);
         #iIndex:= #iIndex+UDINT_TO_UINT(#iTemp3);

         (*Add codeType*)
         Strg_TO_Chars(Strg:= '" codeType="', pChars:= #iIndex, Cnt=> #iTemp3, Chars:=#arrCommand);
         #iIndex:= #iIndex+UDINT_TO_UINT(#iTemp3);
         IF #Data.Matchcode.nCodeType = '*' THEN
           Strg_TO_Chars(Strg:= 'dontCare', pChars:= #iIndex, Cnt=> #iTemp3, Chars:=#arrCommand);
           #iIndex:= #iIndex+UDINT_TO_UINT(#iTemp3);
         ELSE
           #arrCommand[#iIndex]:= #Data.Matchcode.nCodeType;
           #iIndex:= #iIndex+1;
         END_IF;

         (*Add Min/Max length*)
         Strg_TO_Chars(Strg:= '" length="', pChars:= #iIndex, Cnt=> #iTemp3, Chars:=#arrCommand);
         #iIndex:= #iIndex+UDINT_TO_UINT(#iTemp3);
         IF #Data.Matchcode.iMinMaxLength = 0 THEN
           Strg_TO_Chars(Strg:= 'dontCare', pChars:= #iIndex, Cnt=> #iTemp3, Chars:=#arrCommand);
           #iIndex:= #iIndex+UDINT_TO_UINT(#iTemp3);
         ELSE
           #arrCommand[#iIndex]:= ((#Data.Matchcode.iMinMaxLength/100) MOD 10)+16#30;     
           #arrCommand[#iIndex+1]:= ((#Data.Matchcode.iMinMaxLength/10) MOD 10)+16#30;
           #arrCommand[#iIndex+2]:= (#Data.Matchcode.iMinMaxLength MOD 10)+16#30;
           #iIndex:= #iIndex+3;
         END_IF;

         (*Add content*)
         Strg_TO_Chars(Strg:= CONCAT(IN1:= '" content="', IN2:= #Data.Matchcode.sContent), pChars:= #iIndex, Cnt=> #iTemp3, Chars:=#arrCommand);
         #iIndex:= #iIndex+UDINT_TO_UINT(#iTemp3);
         #arrCommand[#iIndex]:= '"';


         (*Overwrite the matchcode length*)
         IF #bCanActive THEN
           #nFncValue:= #iIndex-33;      (*Length of the #Matchcode command*)
           #iCommandLength:= #iIndex+1;  (*Length of the whole CoLa command*)
           #iIndex:= 31;                 (*Startindex of the matchcode length*)
         ELSE
           #nFncValue:= #iIndex-22;      (*Length of the #Matchcode command*)
           #iCommandLength:= #iIndex+1;  (*Length of the whole CoLa command*)
           #iIndex:= 20;                 (*Startindex of the matchcode length*)
         END_IF;

         "SICK_SetValue"(bAddBlank:= false,
                         nValue:= #nFncValue,
                         arrData=> #arrCommand,
                         nErrorCode=> #nFncErrorCode,
                         iPosition:=#iIndex);
         IF #nFncErrorCode <> 16#0000 THEN
           #nTempErrorCode.%W1:= #nFncErrorCode;
           #nTempErrorCode.%W0:= 16#0013; (*Error: SICK_SetValue error*)
         ELSE
           #iStep:= 5; (*Send command*)
         END_IF;

     (*Create "Save Permanent" command*)   
     3:  IF #bCanActive THEN
           Strg_TO_Chars(Strg:= 'MN mEEwriteall', pChars:= 12, Cnt=> #iTemp3, Chars:=#arrCommand);
           #iCommandLength:= UDINT_TO_UINT(#iTemp3+12);
         ELSE
           Strg_TO_Chars(Strg:= 'sMN mEEwriteall', pChars:= 0, Cnt=> #iTemp3, Chars:=#arrCommand);
           #iCommandLength:= UDINT_TO_UINT(#iTemp3);
         END_IF;
         #iStep:= 5; (*Send command*)

     (*Create "Communication Test" command*)
     4:  IF #bCanActive THEN
           Strg_TO_Chars(Strg:= 'RI0', pChars:= 12, Cnt=> #iTemp3, Chars:=#arrCommand);
           #iCommandLength:= UDINT_TO_UINT(#iTemp3)+12;
         ELSE
           Strg_TO_Chars(Strg:= 'sRI0', pChars:= 0, Cnt=> #iTemp3, Chars:=#arrCommand);
           #iCommandLength:= UDINT_TO_UINT(#iTemp3);
         END_IF;
         #iStep:= 5; (*Send command*)

     (*Create "Free Command"*)
     5:  IF #bCanActive THEN
           Strg_TO_Chars(Strg:= DELETE(IN:= #Data.FreeCommand.sCommand, L:=1, P:=1), pChars:= 12, Cnt=> #iTemp3, Chars:=#arrCommand);
           #iCommandLength:= UDINT_TO_UINT(#iTemp3)+12;
         ELSE
           Strg_TO_Chars(Strg:= #Data.FreeCommand.sCommand, pChars:= 0, Cnt=> #iTemp3, Chars:=#arrCommand);
           #iCommandLength:= UDINT_TO_UINT(#iTemp3);
         END_IF;
         #iStep:= 5; (*Send command*)

     (*Create "Login" command*)
     10: IF #bCanActive THEN
           Strg_TO_Chars(Strg:= 'MN SetAccessMode 03 F4724744', pChars:= 12, Cnt=> #iTemp3, Chars:=#arrCommand);
           #iCommandLength:= UDINT_TO_UINT(#iTemp3)+12;
         ELSE
           Strg_TO_Chars(Strg:= 'sMN SetAccessMode 03 F4724744', pChars:= 0, Cnt=> #iTemp3, Chars:=#arrCommand);
           #iCommandLength:= UDINT_TO_UINT(#iTemp3);
         END_IF;
         #iStep:= 5; (*Send command*)

     (*Create "Logout" command*)
     11: IF #bCanActive THEN
           Strg_TO_Chars(Strg:= 'MN Run', pChars:= 12, Cnt=> #iTemp3, Chars:=#arrCommand);
           #iCommandLength:= UDINT_TO_UINT(#iTemp3)+12;
         ELSE
           Strg_TO_Chars(Strg:= 'sMN Run', pChars:= 0, Cnt=> #iTemp3, Chars:=#arrCommand);
           #iCommandLength:= UDINT_TO_UINT(#iTemp3);
         END_IF;
         #iStep:= 5; (*Send command*)

       END_CASE;
   END_IF;


   (*=============================== SEND COLA COMMAND (STEP 5) ===============================*)
   IF #iStep =5 THEN
     IF NOT #fbCCom.ReqBusy AND NOT #bTriggerDone AND NOT #bTriggerError THEN
       #fbCCom.Req:= true;
       #iStep:= 6; (*Wait for the command answer*)
     END_IF;
   END_IF;


   (*========================== WAIT FOR THE COMMAND ANSWER (STEP 6) ==========================*)
   IF #iStep =6 THEN
     (*Communication error*)
     IF #bTriggerError THEN
       #nTempErrorCode:= #fbCCom.Errorcode; (*Error: Communication error*)

       (*Communication done*)
     ELSIF #bTriggerDone THEN
       #iStep:= 7; (*Check the command answer*)
     END_IF;
   END_IF;


   (*============================= CHECK COMMAND RESPONSE (STEP 7) ============================*)
   IF #iStep =7 THEN
     CASE #iCommandIndex OF

     (*Check "Trigger On" response*)
     0:  IF #bCanActive THEN
           IF #arrRecord[0] = 's' AND
             #arrRecord[12] = 'A' AND
             #arrRecord[13] = 'N' AND
             #arrRecord[22] = 'o' AND
             #arrRecord[23] = 'n' AND
             #arrRecord[24] = ' ' AND
             #arrRecord[25] = '1' THEN

             #iStep:= 8; (*Action performed*)
           ELSE
             #nTempErrorCode:= 16#0000_0016; (*Error: Invalid device answer*)                    
           END_IF;
         ELSE
           IF #arrRecord[0] = 's' AND
             #arrRecord[1] = 'A' AND
             #arrRecord[2] = 'N' AND
             #arrRecord[11] = 'o' AND
             #arrRecord[12] = 'n' AND
             #arrRecord[13] = ' ' AND
             #arrRecord[14] = '1' THEN

             #iStep:= 8; (*Action performed*)
           ELSE
             #nTempErrorCode:= 16#0000_0016; (*Error: Invalid device answer*)        
           END_IF;
         END_IF;

     (*Check "Trigger Off" response*)
     1:  IF #bCanActive THEN
           IF #arrRecord[0] = 's' AND
             #arrRecord[12] = 'A' AND
             #arrRecord[13] = 'N' AND
             #arrRecord[22] = 'o' AND
             #arrRecord[23] = 'f' AND
             #arrRecord[24] = 'f' AND
             #arrRecord[25] = ' ' AND
             #arrRecord[26] = '1' THEN

             #iStep:= 8; (*Action performed*)
           ELSE
             #nTempErrorCode:= 16#0000_0016; (*Error: Invalid device answer*)          
           END_IF;
         ELSE
           IF #arrRecord[0] = 's' AND
             #arrRecord[1] = 'A' AND
             #arrRecord[2] = 'N' AND
             #arrRecord[11] = 'o' AND
             #arrRecord[12] = 'f' AND
             #arrRecord[13] = 'f' AND
             #arrRecord[14] = ' ' AND
             #arrRecord[15] = '1' THEN

             #iStep:= 8; (*Action performed*)
           ELSE  
             #nTempErrorCode:= 16#0000_0016; (*Error: Invalid device answer*)          
           END_IF;
         END_IF;

     (*Check "Matchcode" response*)
     2:  IF #bCanActive THEN
           IF NOT(#arrRecord[0] = 's' AND
             #arrRecord[12] = 'A' AND
             #arrRecord[13] = 'N' AND
             #arrRecord[27] = 'o' AND
             #arrRecord[28] = 'd' AND
             #arrRecord[29] = 'e' AND
             #arrRecord[30] = ' ' AND
             #arrRecord[31] = '1') THEN

             #nTempErrorCode:= 16#0000_0016; (*Error: Invalid device answer*)          
           END_IF;
         ELSE
           IF NOT(#arrRecord[0] = 's' AND
             #arrRecord[1] = 'A' AND
             #arrRecord[2] = 'N' AND
             #arrRecord[16] = 'o' AND
             #arrRecord[17] = 'd' AND
             #arrRecord[18] = 'e' AND
             #arrRecord[19] = ' ' AND
             #arrRecord[20] = '1') THEN

             #nTempErrorCode:= 16#0000_0016; (*Error: Invalid device answer*)          
           END_IF;
         END_IF;

         IF #nTempErrorCode = 0 THEN
           #iCommandIndex:= 11; (*Logout*)
           #iStep:= 4;         (*Create command*)
         END_IF;    

     (*Check "Save Permanent" response*)
     3:  IF #bCanActive THEN
           IF NOT(#arrRecord[0] = 's' AND
             #arrRecord[12] = 'A' AND
             #arrRecord[13] = 'N' AND
             #arrRecord[23] = 'a' AND
             #arrRecord[24] = 'l' AND
             #arrRecord[25] = 'l' AND
             #arrRecord[26] = ' ' AND
             #arrRecord[27] = '1') THEN

             #nTempErrorCode:= 16#0000_0016; (*Error: Invalid device answer*)          
           END_IF;
         ELSE
           IF NOT(#arrRecord[0] = 's' AND
             #arrRecord[1] = 'A' AND
             #arrRecord[2] = 'N' AND
             #arrRecord[12] = 'a' AND
             #arrRecord[13] = 'l' AND
             #arrRecord[14] = 'l' AND
             #arrRecord[15] = ' ' AND
             #arrRecord[16] = '1') THEN

             #nTempErrorCode:= 16#0000_0016; (*Error: Invalid device answer*)          
           END_IF;
         END_IF;

         IF #nTempErrorCode = 0 THEN
           #iCommandIndex:= 11; (*Logout*)
           #iStep:= 4;         (*Create command*)
         END_IF;

     (*Check "Communication Test" response*)
     4:  IF #bCanActive THEN
           IF #arrRecord[0] = 's' AND
             #arrRecord[12] = 'R' AND
             #arrRecord[13] = 'A' AND
             #arrRecord[14] = ' ' THEN

             #iStep:= 8; (*Action performed*)
           ELSE
             #nTempErrorCode:= 16#0000_0016; (*Error: Invalid device answer*)          
           END_IF;
         ELSE
           IF #arrRecord[0] = 's' AND
             #arrRecord[1] = 'R' AND
             #arrRecord[2] = 'A' AND
             #arrRecord[3] = ' ' THEN

             #iStep:= 8; (*Action performed*)
           ELSE  
             #nTempErrorCode:= 16#0000_0016; (*Error: Invalid device answer*)          
           END_IF;
         END_IF;

     (*Check "Free command" response*)
     5:  IF #fbCCom.ReqLength <= MAX_LEN(#Data.FreeCommand.sResult) THEN 
           Chars_TO_Strg(Chars:= #arrRecord, pChars:= 0, Cnt:= INT_TO_UINT(#fbCCom.ReqLength),Strg=> #Data.FreeCommand.sResult);
           #iStep:= 8; (*Action performed*)
         ELSE
           #nTempErrorCode:= 16#0000_0021; (*Error: Free command result > Result string*)
         END_IF;

     (*Check "Login" response*)
     10:  IF #bCanActive THEN
           IF NOT(#arrRecord[0] = 's' AND
             #arrRecord[12] = 'A' AND
             #arrRecord[13] = 'N' AND
             #arrRecord[24] = 'M' AND
             #arrRecord[25] = 'o' AND
             #arrRecord[26] = 'd' AND
             #arrRecord[27] = 'e' AND
             #arrRecord[28] = ' ' AND
             #arrRecord[29] = '1') THEN

             #nTempErrorCode:= 16#0000_0016; (*Error: Invalid device answer*)          
           END_IF;
         ELSE
           IF NOT(#arrRecord[0] = 's' AND
             #arrRecord[1] = 'A' AND
             #arrRecord[2] = 'N' AND
             #arrRecord[13] = 'M' AND
             #arrRecord[14] = 'o' AND
             #arrRecord[15] = 'd' AND
             #arrRecord[16] = 'e' AND
             #arrRecord[17] = ' ' AND
             #arrRecord[18] = '1') THEN

             #nTempErrorCode:= 16#0000_0016; (*Error: Invalid device answer*)          
           END_IF;
         END_IF;

         IF #nTempErrorCode = 0 THEN
           IF #arrSelection[2] THEN
             #iCommandIndex:= 2; (*Matchcode*)
             #iStep:= 4;         (*Create command*)
           ELSIF #arrSelection[3] THEN
             #iCommandIndex:= 3; (*Save permanent*)
             #iStep:= 4;         (*Create command*)       
           END_IF;
           #bDeviceState:= true; (*Edit-Mode active*)
         END_IF;

     (*Check "Logout" response*)
     11:  IF #bCanActive THEN
           IF #arrRecord[0] = 's' AND
             #arrRecord[12] = 'A' AND
             #arrRecord[13] = 'N' AND
             #arrRecord[14] = ' ' AND
             #arrRecord[15] = 'R' AND
             #arrRecord[16] = 'u' AND
             #arrRecord[17] = 'n' AND
             #arrRecord[18] = ' ' AND
             #arrRecord[19] = '1' THEN

             #bDeviceState:= false; (*Run-Mode active*)
             #iStep:= 8; (*Action performed*)
           ELSE
             #nTempErrorCode:= 16#0000_0016; (*Error: Invalid device answer*)          
           END_IF;
         ELSE
           IF #arrRecord[0] = 's' AND
             #arrRecord[1] = 'A' AND
             #arrRecord[2] = 'N' AND
             #arrRecord[3] = ' ' AND
             #arrRecord[4] = 'R' AND
             #arrRecord[5] = 'u' AND
             #arrRecord[6] = 'n' AND
             #arrRecord[7] = ' ' AND
             #arrRecord[8] = '1' THEN

             #bDeviceState:= false; (*Run-Mode active*)
             #iStep:= 8; (*Action performed*)
           ELSE  
             #nTempErrorCode:= 16#0000_0016; (*Error: Invalid device answer*)          
           END_IF;
         END_IF;
     END_CASE;
   END_IF;


   (*================================ ACTION PERFORMED (STEP 8) ===============================*)
   IF #iStep =8 THEN
     IF #bEnforceLogout THEN
       #nTempErrorCode:= #nLogoutErrorCode;
     ELSE
       #ReqDone:= true;
       #ReqBusy:= false;
       #bReqBusyMem:= false;
       #iStep:= 0;
     END_IF;
   END_IF;


   (*====================================== COMMUNICATION =====================================*)
   #fbCCom(HWInputIdent:= #HWInputIdent,
           HWInputLength:= #HWInputLength,
           HWOutputIdent:= #HWOutputIdent,
           HWOutputLength:= #HWOutputLength,
           TOut:= #TOut+T#1s,
           CommandLength:= #iCommandLength,
           arrCommand:= #arrCommand,
           arrRecord:= #arrRecord);

   (*Reset the request flag every cycle*)
   #fbCCom.Req:= false;

   (*Read result error*)
   IF #fbCCom.RdLength <0 AND #fbCCom.RdDone THEN
     #Data.ReadingResult.iLength:= -1; (*Error: Reading result longer than record array*)
     FOR #iTemp1:= 1 TO UINT_TO_INT(#iReadingResultSize) DO
       #Data.ReadingResult.arrResult[#iTemp1]:= 16#00;
     END_FOR;

   (*Handling of the reading result*)
   ELSIF #fbCCom.RdDone THEN
     IF #fbCCom.RdLength > #iReadingResultSize THEN
       #Data.ReadingResult.iLength:= -1; (*Error: Reading result longer than reading result array*)
       FOR #iTemp1:= 1 TO UINT_TO_INT(#iReadingResultSize) DO
         #Data.ReadingResult.arrResult[#iTemp1]:= 16#00;
       END_FOR;
     ELSE
       MOVE_BLK(IN:= #arrRecord[0], COUNT:= INT_TO_UINT(#fbCCom.RdLength), OUT=> #Data.ReadingResult.arrResult[1]);
       IF (#Data.ReadingResult.iCounter >=255) THEN
         #Data.ReadingResult.iCounter:= 0;
       ELSE
         #Data.ReadingResult.iCounter:= #Data.ReadingResult.iCounter+1;
       END_IF;
       #Data.ReadingResult.iLength:= #fbCCom.RdLength;
       #RdDone:= true;
     END_IF;
   END_IF;
END_FUNCTION_BLOCK

// folder: SICK AG/Internal

FUNCTION_BLOCK "SICK_CCOMM_PNDP"   // FB10, SCL
TITLE = SICK_CCOM_PNDP / SICK CoLa communication block for AutoIdent devices
{ S7_Optimized_Access := 'TRUE' }
AUTHOR : SICKAG
FAMILY : Ident